(* Logix 5000 project; controller PLC_MCC1201_220AP1 vendor 1 type 14 code 164 rev 35.11; software revision 35.00; part 15 of 25 *)
(* tags used below, declared in another part *)
   AFI : ALIAS FOR B3[7].15;
   AMAX_LEHR_SPD : ALIAS FOR I[81];
   APC_HOST_PERM : ALIAS FOR B3[0].7;
   B3 : DINT[102];
   C5 : COUNTER[100];
   CB_AT_SS_CUTTERS : ALIAS FOR B3[4].0;
   CR1_DOWN_PROX : ALIAS FOR I[64].11;
   CURR_LSD : ALIAS FOR N42[74];
   CURR_MSD : ALIAS FOR N42[73];
   CURR_SYNC : ALIAS FOR N7[2];
   DISTANCE : ALIAS FOR N7[1];
   F96 : REAL[50];
   FLAW_HEAD : ALIAS FOR N43[200];
   FLAW_LANE : ALIAS FOR N43[201];
   FLAW_OFF : ALIAS FOR N43[202];
   FLAW_OUT : ALIAS FOR N7[5];
   FLAW_POS : ALIAS FOR N7[4];
   FLAW_QUEUE : ALIAS FOR N7[9];
   FLAW_XLAT : ALIAS FOR N7[6];
   FLOW_CLK_LSD : ALIAS FOR N7[10];
   FLOW_CLK_MSD : ALIAS FOR N7[11];
   GOOD_FLAW : ALIAS FOR B3[0].0;
   GUN_INDEX : ALIAS FOR N7[0];
   I : INT[128];
   INDEX : ALIAS FOR S[24];
   LEHRSPD_AUTOMAX : ALIAS FOR N98[1];
   LEHRSPD_AVE : ALIAS FOR N98[2];
   LEHRSPD_CURRENT : ALIAS FOR N98[5];
   LEHRSPD_STD : ALIAS FOR N98[3];
   M1_ALM_RESET : ALIAS FOR I[64].9;
   MB_ALM_RESET : ALIAS FOR I[16].10;
   MG59_000 : MESSAGE;   // PIF Operations Write current Lehr speed from N98.5 to N10:10 @ M5
   MG59_002 : MESSAGE;   // PIF Operations Write block N98:0 -> N98:3 to processor M5 N10:16 ->N10:19
   N10 : DINT[128];
   N100 : DINT[1000];
   N11 : DINT[1000];
   N14 : DINT[1000];
   N17 : DINT[1000];
   N20 : DINT[1000];
   N23 : DINT[1000];
   N26 : DINT[1000];
   N29 : DINT[1000];
   N32 : DINT[1000];
   N35 : DINT[1000];
   N38 : DINT[1000];
   N42 : DINT[89];
   N43 : DINT[240];
   N44 : DINT[213];
   N53 : DINT[10];
   N54 : DINT[501];
   N60 : DINT[420];
   N7 : DINT[250];
   N9 : DINT[20];
   N98 : DINT[20];
   N99 : DINT[1000];
   NEXT_SYNC : ALIAS FOR N7[3];
   O : INT[128];
   R97 : CONTROL[4];
   REG_INDEX : DINT;
   REL_CAP_REQUEST : ALIAS FOR I[17].14;
   S : INT[128];
   SPRAY_LENGTH : ALIAS FOR N7[8];
   Status : INT;   // INT tag to retrieve Status value through GSV created during conversion
   T4 : TIMER[100];
   T95 : TIMER[2];
   TMP_d : DINT;
   TMP_xAlwaysOFF : BOOL;
   VHSC_BTR : ALIAS FOR BT41_000;
   VHSC_BTR_E : ALIAS FOR BT41_000.EN;
   VHSC_BTW : ALIAS FOR BT41_001;
   VHSC_CNFG : ALIAS FOR N42[71].0;
   VHSC_WR_EN : ALIAS FOR BT41_001.EN;
(* MainProgram, continued *)

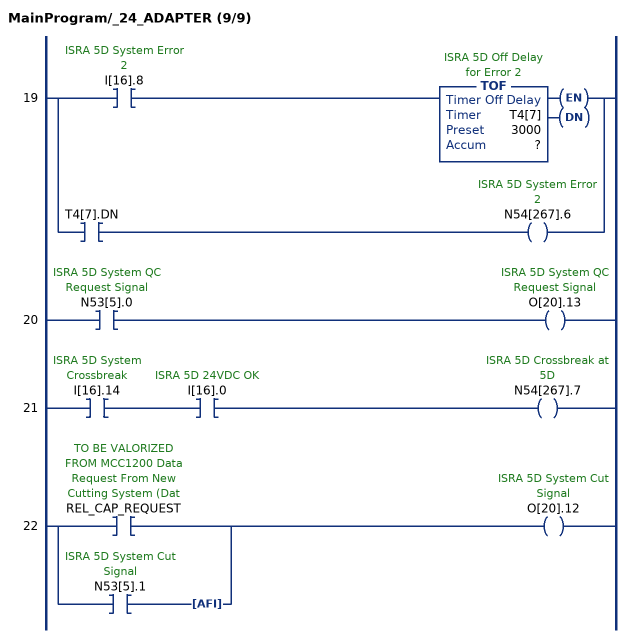
   [picture p214: MainProgram/_24_ADAPTER rungs 19-22]
   19: [XIC(I[16].8) TOF(T4[7],?,?) ,XIC(T4[7].DN) OTE(N54[267].6) ];
   20: XIC(N53[5].0)OTE(O[20].13);
   21: XIC(I[16].14)XIC(I[16].0)OTE(N54[267].7);
   22: [XIC(REL_CAP_REQUEST) ,XIC(N53[5].1) AFI() ]OTE(O[20].12);
END_ROUTINE

ROUTINE _25_PIF_OPS   (* ladder *)
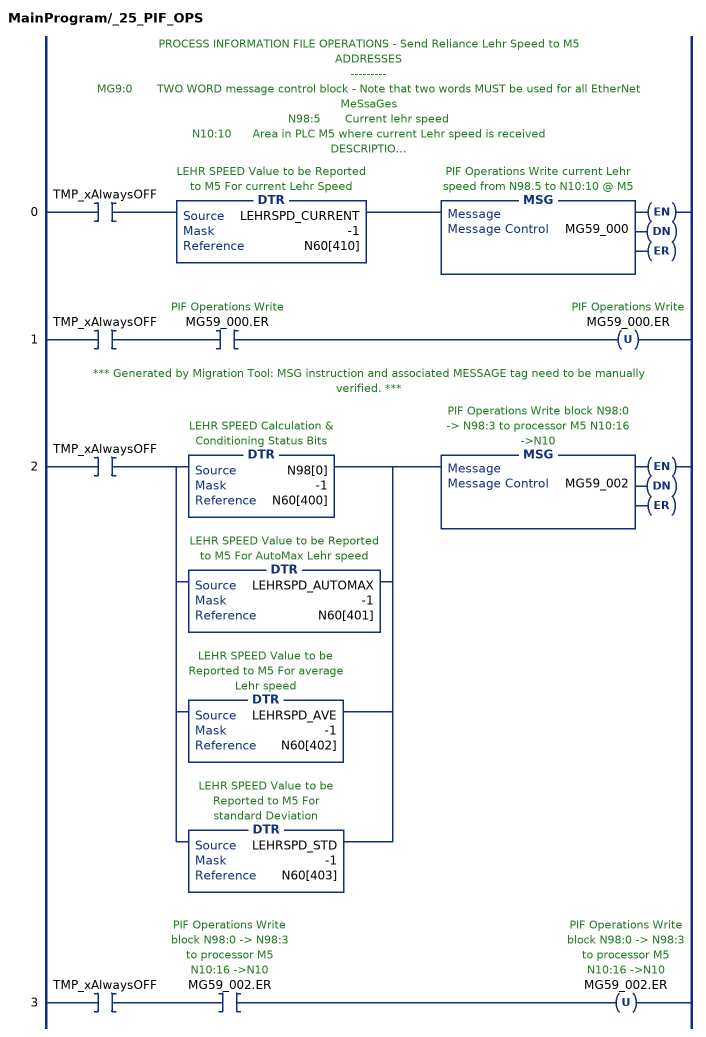
   // PROCESS INFORMATION FILE OPERATIONS - Send Reliance Lehr Speed to M5
   // ADDRESSES
   // ---------
   // MG9:0       TWO WORD message control block - Note that two words MUST be used for all EtherNet MeSsaGes
   // N98:5       Current lehr speed
   // N10:10      Area in PLC M5 where current Lehr speed is received
   // DESCRIPTION
   // -----------
   // This rung transmitts current lehr speed to PLC M5.
   // HISTORY
   // -------
   // DATE        DESCRIPTION                                               PROGRAMMER
   // ----        -----------                                               ----------
   // 4/17/       Enetered rung and comment.                                WAS
   // *** Generated by Migration Tool: MSG instruction and associated MESSAGE tag need to be manually verified. ***
   0: XIC(TMP_xAlwaysOFF)DTR(LEHRSPD_CURRENT,-1,N60[410])MSG(MG59_000);
   1: XIC(TMP_xAlwaysOFF)XIC(MG59_000.ER)OTU(MG59_000.ER);
   // *** Generated by Migration Tool: MSG instruction and associated MESSAGE tag need to be manually verified. ***
   2: XIC(TMP_xAlwaysOFF)[DTR(N98[0],-1,N60[400]) ,DTR(LEHRSPD_AUTOMAX,-1,N60[401]) ,DTR(LEHRSPD_AVE,-1,N60[402]) ,DTR(LEHRSPD_STD,-1,N60[403]) ]MSG(MG59_002);
   3: XIC(TMP_xAlwaysOFF)XIC(MG59_002.ER)OTU(MG59_002.ER);
END_ROUTINE

ROUTINE _27_LEHR_SPD   (* ladder *)
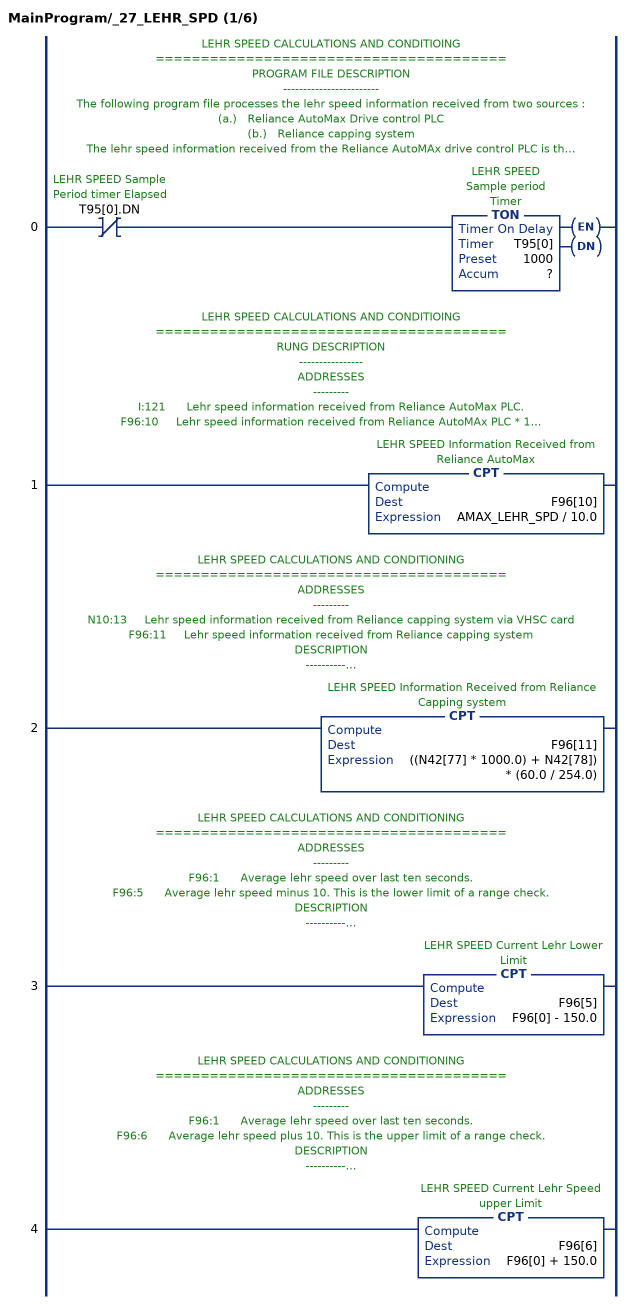
   // LEHR SPEED CALCULATIONS AND CONDITIOING
   // =======================================
   // PROGRAM FILE DESCRIPTION
   // ------------------------
   // The following program file processes the lehr speed information received from two sources :
   //             (a.)   Reliance AutoMax Drive control PLC
   //             (b.)   Reliance capping system
   // The lehr speed information received from the Reliance AutoMAx drive control PLC is the primary
   // source of lehr speed. If this is determined to be invalid, the the data received from the Reliance
   // capping system is used. If neither sourse contains valid data, then the average lehr speed over
   // the last ten seconds is used.
   // The lehr speed can be reset by pressing the "alarm reset" pushbutton located at the No. 1 crusher panel
   // or on VMCC M2.
   // RUNG DESCRIPTION
   // ----------------
   // This rung drives a sample period timer. The timer duration is 1 second.
   // HISTORY
   // DATE        DESCRIPTION                                                  PROGRAMMER
   // ====        ===========                                                  ==========
   // 4/17/96     Entered rungs and comments                                   WAS
   0: XIO(T95[0].DN)TON(T95[0],?,?);
   // LEHR SPEED CALCULATIONS AND CONDITIOING
   // =======================================
   // RUNG DESCRIPTION
   // ----------------
   // ADDRESSES
   // ---------
   // I:121      Lehr speed information received from Reliance AutoMax PLC.
   // F96:10     Lehr speed information received from Reliance AutoMAx PLC * 10
   // DESCRIPTION
   // -----------
   // The data received from the Reliance AutoMax PLC is in the form :
   //           Lehr Speed * 10
   // This rung divides the value received from the AutoMax PLC by 10 and
   // writes it into F96:10.
   // HISTORY
   // DATE        DESCRIPTION                                                  PROGRAMMER
   // ====        ===========                                                  ==========
   // 4/17/96     Entered rungs and comments                                   WAS
   1: CPT(F96[10],AMAX_LEHR_SPD / 10.0);
   // LEHR SPEED CALCULATIONS AND CONDITIONING
   // =======================================
   // ADDRESSES
   // ---------
   // N10:13     Lehr speed information received from Reliance capping system via VHSC card
   // F96:11     Lehr speed information received from Reliance capping system
   // DESCRIPTION
   // -----------
   // The data received from the Reliance capping system is in the form :
   //           1 pulse per 0.1 millimeters of travel
   // The VHSC card receives the 1/10th of a millimeter pulse on VHSC counter 2. It provides a
   // frequency for this pulse train in N42:77 and N42:78, where N42:77 is NNN in NNN,xxx and N42:77
   // is xxx,NNN. The conversion constant is (60/254) is from the following :
   //                1 Pulse     60 sec.       1 in
   //                _______  x  ______     x  _______
   //                0.1 mm      1 min.        254 mm.
   // The resultant conversion constant has an approximate value of 0.2362204724409, and
   // is used to convert the 0.1 mm. pulse to inches per minute.
   // HISTORY
   // DATE        DESCRIPTION                                                  PROGRAMMER
   // ====        ===========                                                  ==========
   // 4/17/96     Entered rungs and comments                                   WAS
   2: CPT(F96[11],((N42[77] * 1000.0) + N42[78]) * (60.0 / 254.0));
   // LEHR SPEED CALCULATIONS AND CONDITIONING
   // =======================================
   // ADDRESSES
   // ---------
   // F96:1      Average lehr speed over last ten seconds.
   // F96:5      Average lehr speed minus 10. This is the lower limit of a range check.
   // DESCRIPTION
   // -----------
   // The rung calculates the lower limit for a range check.
   // HISTORY
   // DATE        DESCRIPTION                                                  PROGRAMMER
   // ====        ===========                                                  ==========
   // 4/17/96     Entered rungs and comments                                   WAS
   3: CPT(F96[5],F96[0] - 150.0);
   // LEHR SPEED CALCULATIONS AND CONDITIONING
   // =======================================
   // ADDRESSES
   // ---------
   // F96:1      Average lehr speed over last ten seconds.
   // F96:6      Average lehr speed plus 10. This is the upper limit of a range check.
   // DESCRIPTION
   // -----------
   // The rung calculates the upper limit for a range check.
   // HISTORY
   // DATE        DESCRIPTION                                                  PROGRAMMER
   // ====        ===========                                                  ==========
   // 4/17/96     Entered rungs and comments                                   WAS
   4: CPT(F96[6],F96[0] + 150.0);
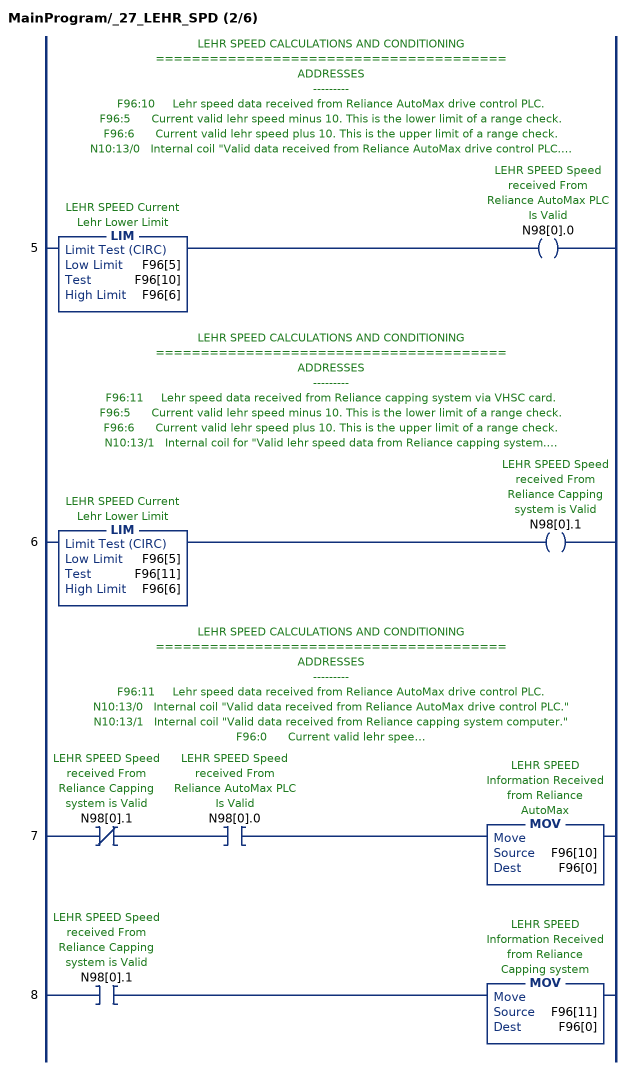
   // LEHR SPEED CALCULATIONS AND CONDITIONING
   // =======================================
   // ADDRESSES
   // ---------
   // F96:10     Lehr speed data received from Reliance AutoMax drive control PLC.
   // F96:5      Current valid lehr speed minus 10. This is the lower limit of a range check.
   // F96:6      Current valid lehr speed plus 10. This is the upper limit of a range check.
   // N10:13/0   Internal coil "Valid data received from Reliance AutoMax drive control PLC."
   // DESCRIPTION
   // -----------
   // This rung determines if the current lehr speed data received from the
   // Reliance AutoMax drive control PLC is valid. The data is compared to a
   // range check with the following limits :
   //             Average Lehr Speed - 10
   //             Average Lehr Speed + 10
   // If the lehr speed is found to be within these limits, then the coil N10:13/0 is set
   // indicating valid lehr speed data from the Reliance AutoMax drive control PLC.
   // HISTORY
   // DATE        DESCRIPTION                                                  PROGRAMMER
   // ====        ===========                                                  ==========
   // 4/17/96     Entered rungs and comments                                   WAS
   5: LIM(F96[5],F96[10],F96[6])OTE(N98[0].0);
   // LEHR SPEED CALCULATIONS AND CONDITIONING
   // =======================================
   // ADDRESSES
   // ---------
   // F96:11     Lehr speed data received from Reliance capping system via VHSC card.
   // F96:5      Current valid lehr speed minus 10. This is the lower limit of a range check.
   // F96:6      Current valid lehr speed plus 10. This is the upper limit of a range check.
   // N10:13/1   Internal coil for "Valid lehr speed data from Reliance capping system."
   // DESCRIPTION
   // -----------
   // This rung determines if the current lehr speed data received from the
   // Reliance capping system is valid. The data is compared to a range check
   //  with the following limits :
   //             Average Lehr Speed - 10
   //             Average Lehr Speed + 10
   // If the lehr speed is found to be within these limits, then the coil N10:13/1 is set
   // indicating valid lehr speed data from the Reliance capping system computer.
   // HISTORY
   // DATE        DESCRIPTION                                                  PROGRAMMER
   // ====        ===========                                                  ==========
   // 4/17/96     Entered rungs and comments                                   WAS
   6: LIM(F96[5],F96[11],F96[6])OTE(N98[0].1);
   // LEHR SPEED CALCULATIONS AND CONDITIONING
   // =======================================
   // ADDRESSES
   // ---------
   // F96:11     Lehr speed data received from Reliance AutoMax drive control PLC.
   // N10:13/0   Internal coil "Valid data received from Reliance AutoMax drive control PLC."
   // N10:13/1   Internal coil "Valid data received from Reliance capping system computer."
   // F96:0      Current valid lehr speed
   // DESCRIPTION
   // -----------
   // If the data from the Reliance AutoMax drive control PLC is NOT valid,
   // but the data from th Reliance capping system IS valid, then it shall
   // be used as the current valid lehr speed.
   // HISTORY
   // DATE        DESCRIPTION                                                  PROGRAMMER
   // ====        ===========                                                  ==========
   // 4/17/96     Entered rungs and comments                                   WAS
   7: XIO(N98[0].1)XIC(N98[0].0)MOV(F96[10],F96[0]);
   8: XIC(N98[0].1)MOV(F96[11],F96[0]);
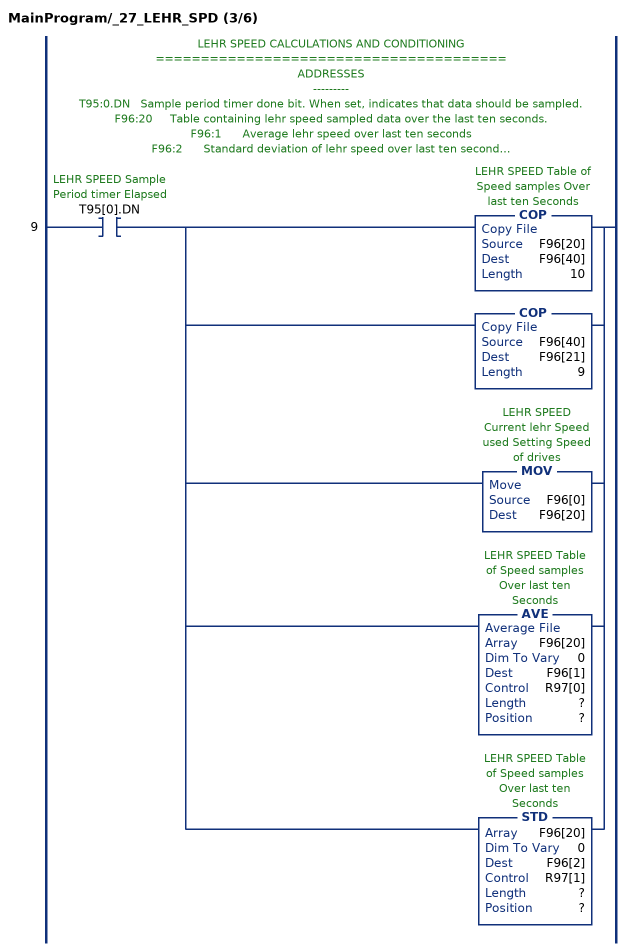
   // LEHR SPEED CALCULATIONS AND CONDITIONING
   // =======================================
   // ADDRESSES
   // ---------
   // T95:0.DN   Sample period timer done bit. When set, indicates that data should be sampled.
   // F96:20     Table containing lehr speed sampled data over the last ten seconds.
   // F96:1      Average lehr speed over last ten seconds
   // F96:2      Standard deviation of lehr speed over last ten seconds
   // F96:0      Current valid lehr speed
   // R97:0      Control file for Average calculation
   // R97:1      Control file for Standard deviation calculation
   // DESCRIPTION
   // -----------
   // When the sample period timer has elapsed, then the stack for lehr speed
   // data over the last ten seconds is updated with the current valid lehr speed.
   // This is accomplished with the COP instruction and MOV instruction.
   // The AVE and STD instructions are used to calcuate the average and standard
   // deviation on the table, respectively.
   // HISTORY
   // DATE        DESCRIPTION                                                  PROGRAMMER
   // ====        ===========                                                  ==========
   // 4/17/96     Entered rungs and comments                                   WAS
   9: XIC(T95[0].DN)[COP(F96[20],F96[40],10) ,COP(F96[40],F96[21],9) ,MOV(F96[0],F96[20]) ,AVE(F96[20],0,F96[1],R97[0],?,?) ,STD(F96[20],0,F96[2],R97[1],?,?) ];
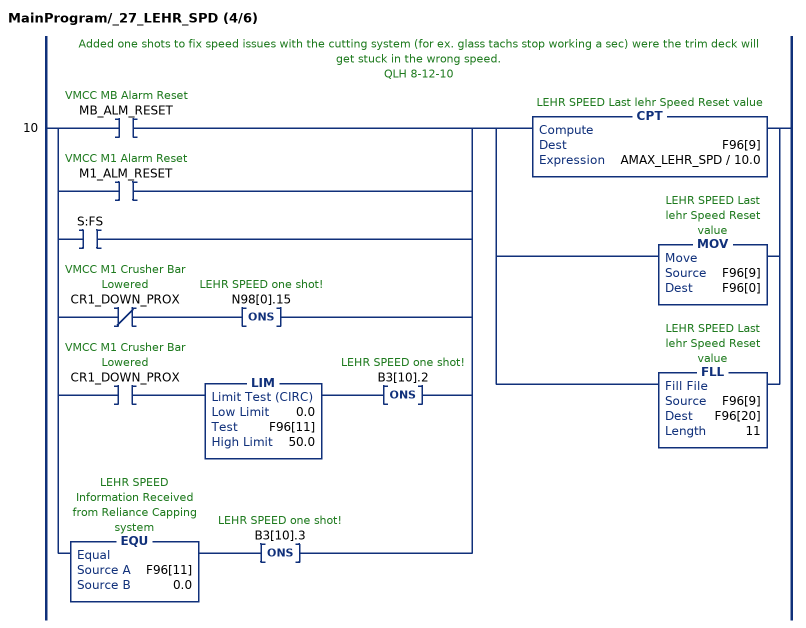
   // Added one shots to fix speed issues with the cutting system (for ex. glass tachs stop working a sec) were the trim deck will get stuck in the wrong speed.
   // QLH 8-12-10
   10: [XIC(MB_ALM_RESET) ,XIC(M1_ALM_RESET) ,XIC(S:FS) ,XIO(CR1_DOWN_PROX) ONS(N98[0].15) ,XIC(CR1_DOWN_PROX) LIM(0.0,F96[11],50.0) ONS(B3[10].2) ,EQU(F96[11],0.0) ONS(B3[10].3) ][CPT(F96[9],AMAX_LEHR_SPD / 10.0) ,MOV(F96[9],F96[0]) ,FLL(F96[9],F96[20],11) ];
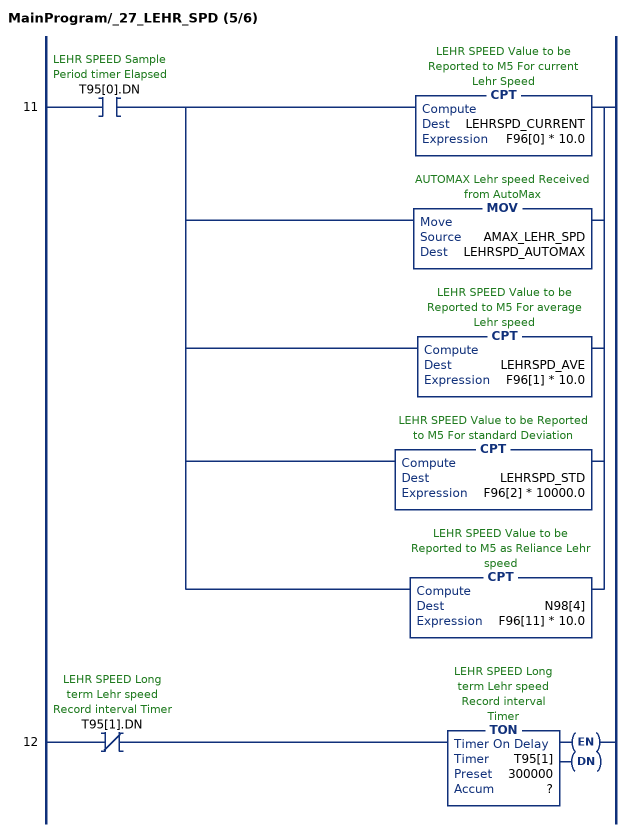
   11: XIC(T95[0].DN)[CPT(LEHRSPD_CURRENT,F96[0] * 10.0) ,MOV(AMAX_LEHR_SPD,LEHRSPD_AUTOMAX) ,CPT(LEHRSPD_AVE,F96[1] * 10.0) ,CPT(LEHRSPD_STD,F96[2] * 10000.0) ,CPT(N98[4],F96[11] * 10.0) ];
   12: XIO(T95[1].DN)TON(T95[1],?,?);
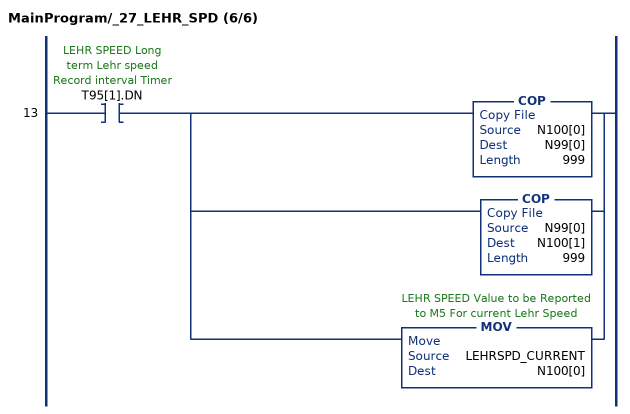
   13: XIC(T95[1].DN)[COP(N100[0],N99[0],999) ,COP(N99[0],N100[1],999) ,MOV(LEHRSPD_CURRENT,N100[0]) ];
END_ROUTINE

ROUTINE _2_TRACKING   (* ladder *)
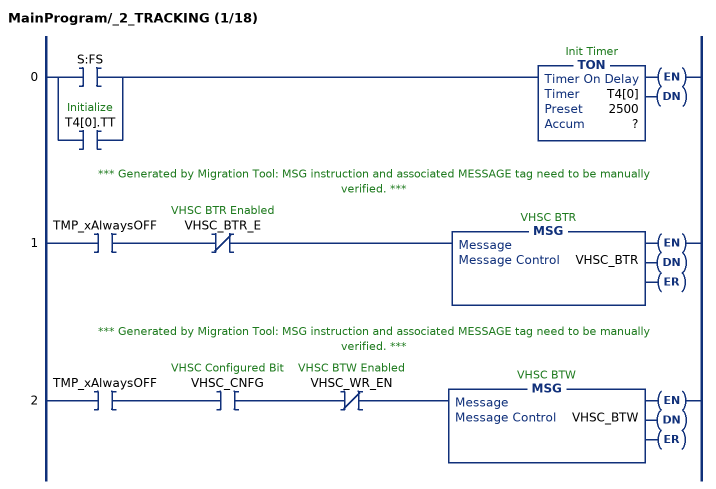
   0: [XIC(S:FS) ,XIC(T4[0].TT) ]TON(T4[0],?,?);
   // *** Generated by Migration Tool: MSG instruction and associated MESSAGE tag need to be manually verified. ***
   1: XIC(TMP_xAlwaysOFF)XIO(VHSC_BTR_E)MSG(VHSC_BTR);
   // *** Generated by Migration Tool: MSG instruction and associated MESSAGE tag need to be manually verified. ***
   2: XIC(TMP_xAlwaysOFF)XIC(VHSC_CNFG)XIO(VHSC_WR_EN)MSG(VHSC_BTW);
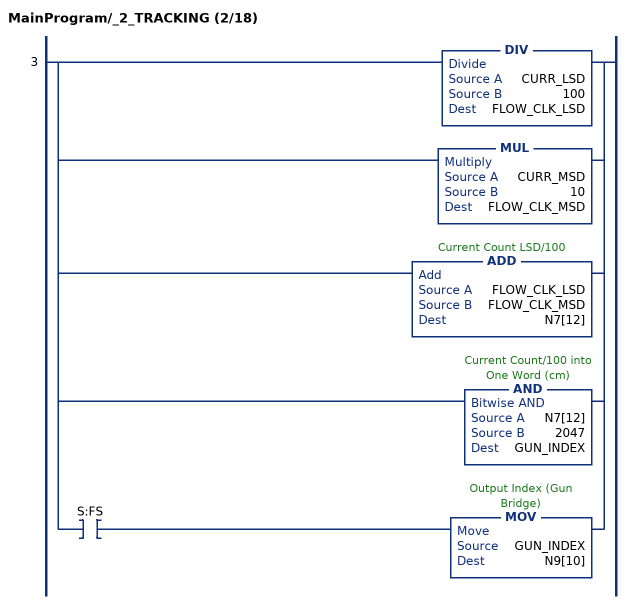
   3: [DIV(CURR_LSD,100,FLOW_CLK_LSD) ,MUL(CURR_MSD,10,FLOW_CLK_MSD) ,ADD(FLOW_CLK_LSD,FLOW_CLK_MSD,N7[12]) ,AND(N7[12],2047,GUN_INDEX) ,XIC(S:FS) MOV(GUN_INDEX,N9[10]) ];
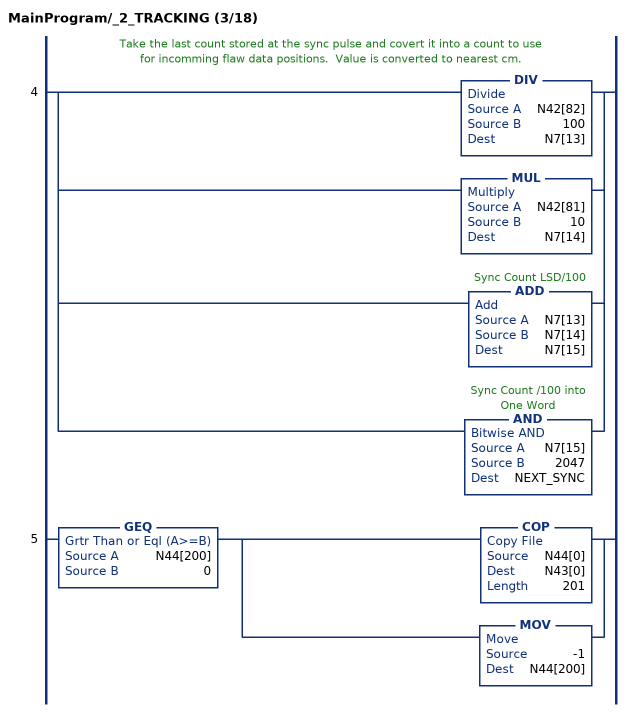
   // Take the last count stored at the sync pulse and covert it into a count to use
   // for incomming flaw data positions.  Value is converted to nearest cm.
   4: [DIV(N42[82],100,N7[13]) ,MUL(N42[81],10,N7[14]) ,ADD(N7[13],N7[14],N7[15]) ,AND(N7[15],2047,NEXT_SYNC) ];
   5: GEQ(N44[200],0)[COP(N44[0],N43[0],201) ,MOV(-1,N44[200]) ];